               x8 : Bool;   // P2648.EPOS direct setpoint input/MDI positioning type
               x9 : Bool;   // P2651.EPOS direct setpoint input/MDI direction selection positive
               x10 : Bool;   // P2652.EPOS direct setpoint input/MDI direction selection negative
               x11 : Bool;   // Reserved
               x12 : Bool;   // P2649.EPOS direct setpoint input/MDI transfer type selection
               x13 : Bool;   // Reserved
               x14 : Bool;   // P2653.EPOS direct setpoint input/MDI setting-up selection
               x15 : Bool;   // P2647.EPOS direct setpoint input/MDI selection
               x0 : Bool;   // P2525.EPOS traversing block selection, bit 0
               x1 : Bool;   // P2526.EPOS traversing block selection, bit 1
               x2 : Bool;   // P2527.EPOS traversing block selection, bit 2
               x3 : Bool;   // P2528.EPOS traversing block selection, bit 3
               x4 : Bool;   // P2529.EPOS traversing block selection, bit 4
               x5 : Bool;   // P2530.EPOS traversing block selection, bit 5
               x6 : Bool;   // Reserved
               x7 : Bool;   // P2577.EPOS module correction activation
            END_STRUCT;
            tPOS_STW2 : Struct   // POSITIONER CONTROL WORD 3
               x8 : Bool;   // P2597.EPOS referencing type selection
               x9 : Bool;   // P2604.EPOS search for reference, start direction
               x10 : Bool;   // P2510.LR selecting measuring probe evaluation
               x11 : Bool;   // P2511.LR measuring probe evaluation edge
               x12 : Bool;   // Reserved
               x13 : Bool;   // Reserved
               x14 : Bool;   // P2582.EPOS software limit switch activation
               x15 : Bool;   // P2568.EPOS STOP cam activation
               x0 : Bool;   // P2655.EPOS select tracking mode
               x1 : Bool;   // P2596.EPOS set reference point
               x2 : Bool;   // P2612.EPOS search for reference cam
               x3 : Bool;   // Reserved
               x4 : Bool;   // Reserved
               x5 : Bool;   // P2591.EPOS jogging incremental
               x6 : Bool;   // Reserved
               x7 : Bool;   // Reserved
            END_STRUCT;
            iSTW2 : Int;   // P2045.CONTROL WORD 4
            iOVERRIDE : Int;   // P2646.Override % [0-16384]
            dMDI_TARPOS : DInt;   // P2642.Target position for MDI
            dMDI_VELOCITY : DInt;   // P2643.Speed reference for MDI
            iMDI_ACC : Int;   // P2644.Acceleration ramp % for MDI [0-16384]
            iMDI_DEC : Int;   // P2645.Deceleration ramp % for MDI [0-16384]
            iUser : Int;
         END_STRUCT;
      END_STRUCT;
   END_VAR
   VAR_TEMP
      TMP_dOldValue_AR1 : DInt;
      TMP_dOldValue_AR2 : DInt;
      TMP_x : Bool;
      TMP_i : Int;
      TMP_d : DInt;
      TMP_r : Real;
      TMP_a : ANY;
      TMP_dZero : DInt;
      TMP_xAlwaysON : Bool;
      TMP_rActualSpeed : Real;
      TMP_iAddressLength : Int;
      TMP_dActualPosMin_dmm : DInt;   // Actual position minimum tollerance [mm/10]
      TMP_dActualPosMax_dmm : DInt;   // Actual position maximum tollerance [mm/10]
      TMP_iRetVal : Int;
   END_VAR
   VAR_TEMP   // added for the SCL form of the ladder/FBD networks
      _w1 : Bool;
      _w2 : Bool;
      _w3 : Bool;
      _w4 : Bool;
      _w5 : Bool;
      _w6 : Bool;
      _w7 : Bool;
      _w8 : Bool;
      _w9 : Bool;
      _w10 : Bool;
      _w11 : Bool;
      _w12 : Bool;
   END_VAR
BEGIN

REGION Network 1 (STL): Save AR1 & AR2 value
   //    TAR1
   //    T     #TMP_dOldValue_AR1
   //    TAR2
   //    T     #TMP_dOldValue_AR2
END_REGION

REGION Network 2: #####_COSTANTS_#####
END_REGION

REGION Network 3 (STL): Initializing
         SET;
         S     #TMP_xAlwaysON;

         L     DINT#0;
         T     #TMP_dZero;

         CALL  FILL
         ( BVAL    := #TMP_dZero,
           RET_VAL := #TMP_iRetVal,
           BLK     := #STC_tPZD_Pos.tR
         );
END_REGION

REGION Network 4: #####_MOTOR_MODULE_#####
END_REGION

REGION Network 5 (STL): Check system data coerence
         L     #STC_tSYS_DATA.iIOAddress_MM;
         L     0;
         <I;
         L     10;
         JC    Err;

         L     #STC_tSYS_DATA.dMaxSpeed_rpm;
         L     DINT#0;
         <=D;
         L     11;
         JC    Err;

         L     #STC_tSYS_DATA.rK_rpm_mmMin;
         L     0.0;
         <=R;
         L     12;
         JC    Err;

         L     #STC_tSYS_DATA.rMaxAcc_m_s2;
         L     0.0;
         <=R;
         L     14;
         JC    Err;

         L     #STC_tSYS_DATA.rMaxDec_m_s2;
         L     0.0;
         <=R;
         L     15;
         JC    Err;

         L     12;
         T     #TMP_iAddressLength;

   //Compute destination position
         L;
         LAR1;
   //byte 1 = 10h (FIXED for S7)
         L     B#16#10;
         T     B[AR1, P#0.0];
   //byte 2 = data type
         L     B#16#4;  //4 = word
         T     B[AR1, P#1.0];
   //byte 3 & 4 = number of element
         L     #TMP_iAddressLength;  //Production data
         T     W[AR1, P#2.0];
   //byte 5 & 6 = number of DB
         L     0;  //DB production data
         T     W[AR1, P#4.0];
   //byte 7 = memory area
         L     B#16#81;  //81h = I (Input)
         T     B[AR1, P#6.0];
   //byte 8 & 9 = address. Bit 0,1,2 of tenth byte is bit offset
   //byte 7 = address (high). Valid value = 0-7. Bit 3,4,5,6,7 always 0

         L     #STC_tSYS_DATA.iIOAddress_MM;  //Item size
         SLW   3;
         T     W[AR1, P#8.0];
         SRD   16;
         AW    16#0007;
         T     B[AR1, P#7.0];

         CALL  BLKMOV
         ( SRCBLK  := #TMP_a,
           RET_VAL := #TMP_iRetVal,
           DSTBLK  := #STC_tPZD_Pos.tR
         );
END_REGION

REGION Network 6: #########################_POSITIONER_###########################
END_REGION

REGION Network 7: #####_MATCH_#####
END_REGION

REGION Network 8: Status signals
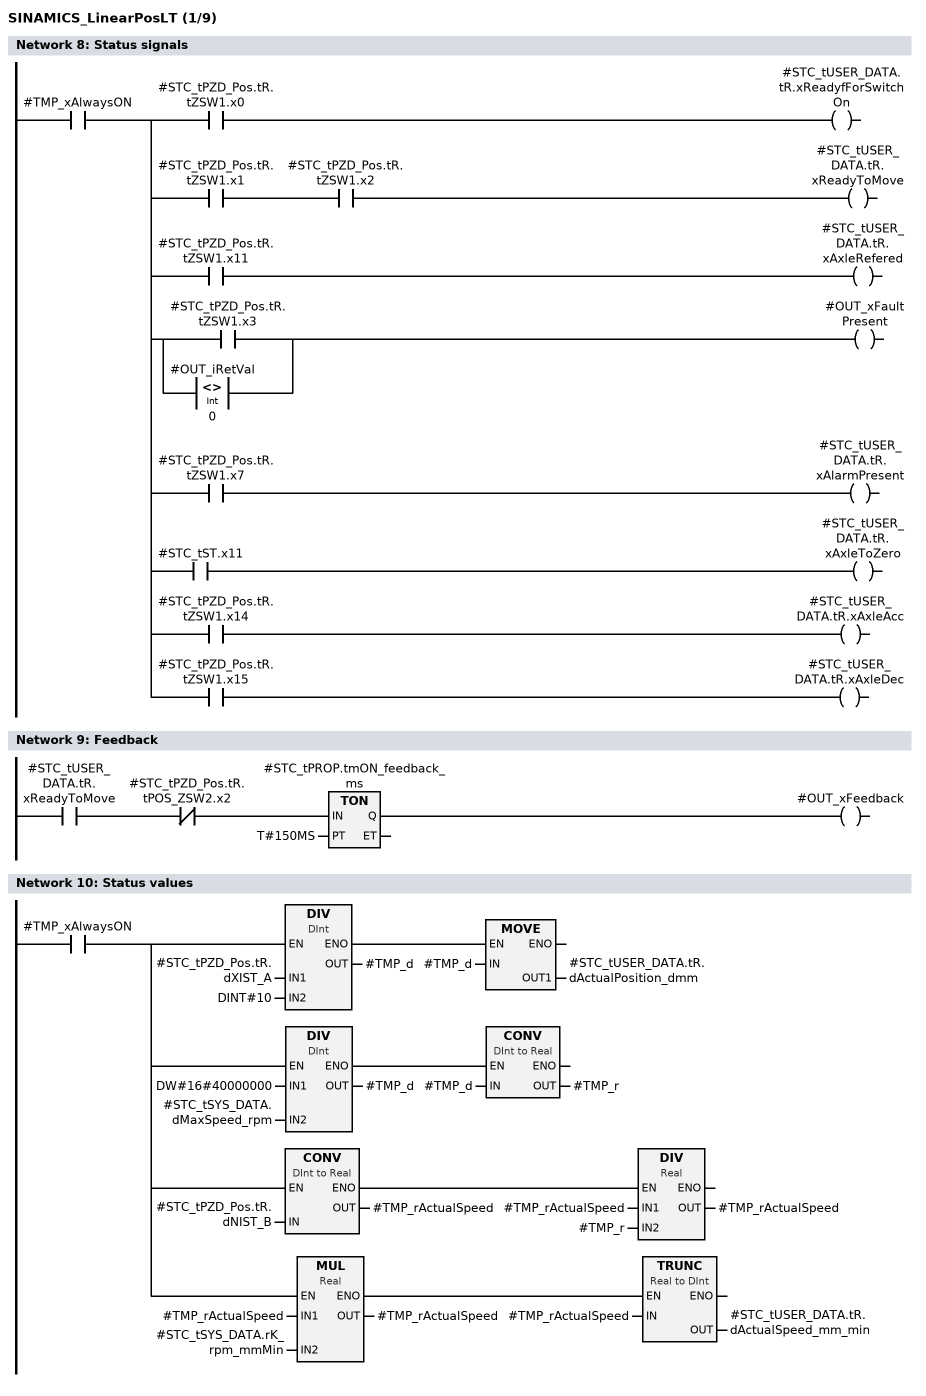
   RUNG wire#powerrail
      Contact( #TMP_xAlwaysON )
      wire#w1
      Contact( #STC_tPZD_Pos.tR.tZSW1.x0 )
      Coil( #STC_tUSER_DATA.tR.xReadyfForSwitchOn )
   END_RUNG
   RUNG wire#w1
      Contact( #STC_tPZD_Pos.tR.tZSW1.x1 )
      Contact( #STC_tPZD_Pos.tR.tZSW1.x2 )
      Coil( #STC_tUSER_DATA.tR.xReadyToMove )
   END_RUNG
   RUNG wire#w1
      Contact( #STC_tPZD_Pos.tR.tZSW1.x11 )
      Coil( #STC_tUSER_DATA.tR.xAxleRefered )
   END_RUNG
   RUNG wire#w1
      Contact( #STC_tPZD_Pos.tR.tZSW1.x3 )
      wire#w2
      Coil( #OUT_xFaultPresent )
   END_RUNG
   RUNG wire#w1
      { S7_Templates := "SrcType := Int" } NE_Contact(in1 := #OUT_iRetVal, in2 := 0)
   END_RUNG wire#w2
   RUNG wire#w1
      Contact( #STC_tPZD_Pos.tR.tZSW1.x7 )
      Coil( #STC_tUSER_DATA.tR.xAlarmPresent )
   END_RUNG
   RUNG wire#w1
      Contact( #STC_tST.x11 )
      Coil( #STC_tUSER_DATA.tR.xAxleToZero )
   END_RUNG
   RUNG wire#w1
      Contact( #STC_tPZD_Pos.tR.tZSW1.x14 )
      Coil( #STC_tUSER_DATA.tR.xAxleAcc )
   END_RUNG
   RUNG wire#w1
      Contact( #STC_tPZD_Pos.tR.tZSW1.x15 )
      Coil( #STC_tUSER_DATA.tR.xAxleDec )
   END_RUNG
   // the same network as SCL:
   #STC_tUSER_DATA.tR.xReadyfForSwitchOn := #TMP_xAlwaysON AND #STC_tPZD_Pos.tR.tZSW1.x0;
   #STC_tUSER_DATA.tR.xReadyToMove := #TMP_xAlwaysON AND #STC_tPZD_Pos.tR.tZSW1.x1 AND #STC_tPZD_Pos.tR.tZSW1.x2;
   #STC_tUSER_DATA.tR.xAxleRefered := #TMP_xAlwaysON AND #STC_tPZD_Pos.tR.tZSW1.x11;
   #OUT_xFaultPresent := #TMP_xAlwaysON AND (#STC_tPZD_Pos.tR.tZSW1.x3 OR (#OUT_iRetVal <> 0));
   #STC_tUSER_DATA.tR.xAlarmPresent := #TMP_xAlwaysON AND #STC_tPZD_Pos.tR.tZSW1.x7;
   #STC_tUSER_DATA.tR.xAxleToZero := #TMP_xAlwaysON AND #STC_tST.x11;
   #STC_tUSER_DATA.tR.xAxleAcc := #TMP_xAlwaysON AND #STC_tPZD_Pos.tR.tZSW1.x14;
   #STC_tUSER_DATA.tR.xAxleDec := #TMP_xAlwaysON AND #STC_tPZD_Pos.tR.tZSW1.x15;
END_REGION

REGION Network 9: Feedback
   #STC_tPROP.tmON_feedback_ms.TON(IN := #STC_tUSER_DATA.tR.xReadyToMove AND NOT #STC_tPZD_Pos.tR.tPOS_ZSW2.x2,
                           PT := T#150MS);
   #OUT_xFeedback := #STC_tPROP.tmON_feedback_ms.Q;
END_REGION

REGION Network 10: Status values
   RUNG wire#powerrail
      Contact( #TMP_xAlwaysON )
      wire#w1
      { S7_Templates := "SrcType := DInt"; S7_GenerateENO := "TRUE" } Div(in1 := #STC_tPZD_Pos.tR.dXIST_A, in2 := DINT#10, out => #TMP_d)
      { S7_GenerateENO := "TRUE" } Move(in := #TMP_d, out1 => #STC_tUSER_DATA.tR.dActualPosition_dmm)
   END_RUNG
   RUNG wire#w1
      { S7_Templates := "SrcType := DInt"; S7_GenerateENO := "TRUE" } Div(in1 := DW#16#40000000, in2 := #STC_tSYS_DATA.dMaxSpeed_rpm, out => #TMP_d)
      { S7_Templates := "[SrcType := DInt, DestType := Real]"; S7_GenerateENO := "TRUE" } Convert(in := #TMP_d, out => #TMP_r)
   END_RUNG
   RUNG wire#w1
      { S7_Templates := "[SrcType := DInt, DestType := Real]"; S7_GenerateENO := "TRUE" } Convert(in := #STC_tPZD_Pos.tR.dNIST_B, out => #TMP_rActualSpeed)
      { S7_Templates := "SrcType := Real"; S7_GenerateENO := "TRUE" } Div(in1 := #TMP_rActualSpeed, in2 := #TMP_r, out => #TMP_rActualSpeed)
   END_RUNG
   RUNG wire#w1
      { S7_Templates := "SrcType := Real"; S7_GenerateENO := "TRUE" } Mul(in1 := #TMP_rActualSpeed, in2 := #STC_tSYS_DATA.rK_rpm_mmMin, out => #TMP_rActualSpeed)
      { S7_Templates := "[SrcType := Real, DestType := DInt]"; S7_GenerateENO := "TRUE" } Trunc(in := #TMP_rActualSpeed, out => #STC_tUSER_DATA.tR.dActualSpeed_mm_min)
   END_RUNG
   // the same network as SCL:
   // ENO of a box is taken as its EN; it also drops when the box reports an error
   IF #TMP_xAlwaysON THEN
       #TMP_d := #STC_tPZD_Pos.tR.dXIST_A / DINT#10;
       #STC_tUSER_DATA.tR.dActualPosition_dmm := #TMP_d;
       #TMP_d := DW#16#40000000 / #STC_tSYS_DATA.dMaxSpeed_rpm;
       #TMP_r := DINT_TO_REAL(#TMP_d);
       #TMP_rActualSpeed := DINT_TO_REAL(#STC_tPZD_Pos.tR.dNIST_B);
       #TMP_rActualSpeed := #TMP_rActualSpeed / #TMP_r;
       #TMP_rActualSpeed := #TMP_rActualSpeed * #STC_tSYS_DATA.rK_rpm_mmMin;
       #STC_tUSER_DATA.tR.dActualSpeed_mm_min := TRUNC(#TMP_rActualSpeed);
   END_IF;
END_REGION

REGION Network 11: #####_STATUSES_#####
END_REGION

REGION Network 12: Type of positioning
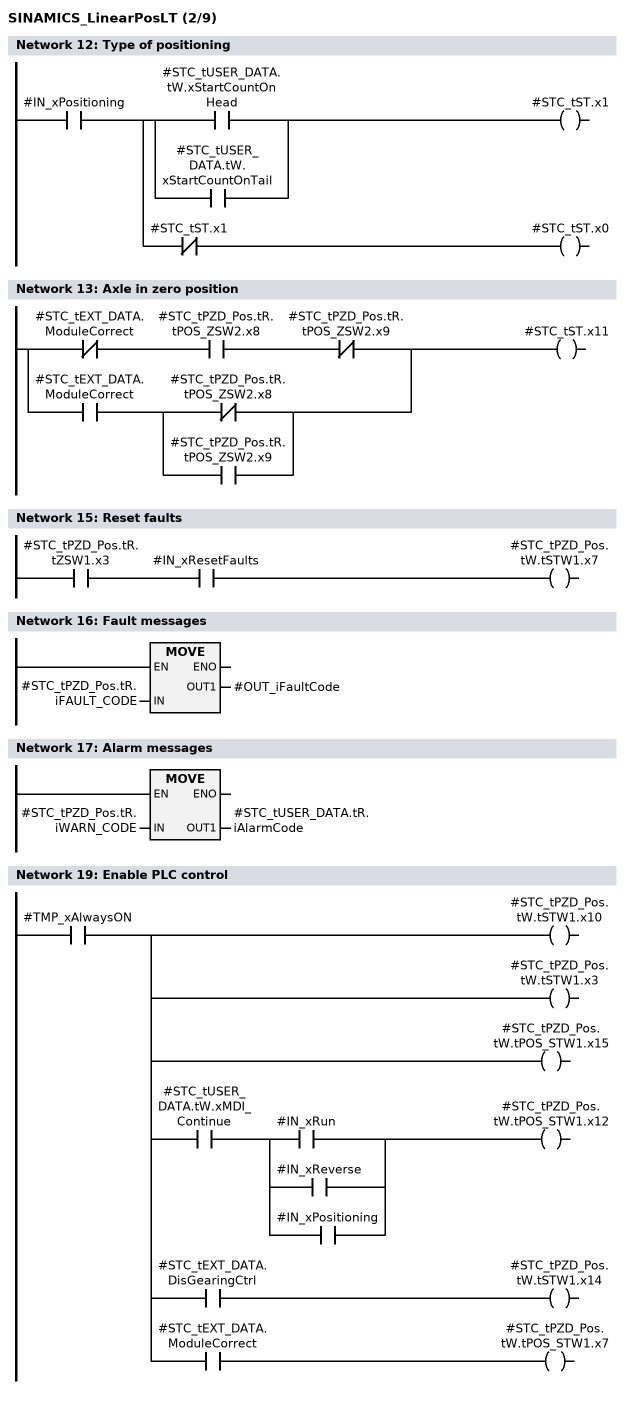
   RUNG wire#powerrail
      Contact( #IN_xPositioning )
      wire#w1
      Contact( #STC_tUSER_DATA.tW.xStartCountOnHead )
      wire#w2
      Coil( #STC_tST.x1 )
   END_RUNG
   RUNG wire#w1
      Contact( #STC_tUSER_DATA.tW.xStartCountOnTail )
   END_RUNG wire#w2
   RUNG wire#w1
      I_Contact( #STC_tST.x1 )
      Coil( #STC_tST.x0 )
   END_RUNG
   // the same network as SCL:
   #STC_tST.x1 := #IN_xPositioning AND (#STC_tUSER_DATA.tW.xStartCountOnHead OR #STC_tUSER_DATA.tW.xStartCountOnTail);
   #STC_tST.x0 := #IN_xPositioning AND NOT #STC_tST.x1;
END_REGION

REGION Network 13: Axle in zero position
   RUNG wire#powerrail
      I_Contact( #STC_tEXT_DATA.ModuleCorrect )
      Contact( #STC_tPZD_Pos.tR.tPOS_ZSW2.x8 )
      I_Contact( #STC_tPZD_Pos.tR.tPOS_ZSW2.x9 )
      wire#w1
      Coil( #STC_tST.x11 )
   END_RUNG
   RUNG wire#powerrail
      Contact( #STC_tEXT_DATA.ModuleCorrect )
      wire#w2
      I_Contact( #STC_tPZD_Pos.tR.tPOS_ZSW2.x8 )
   END_RUNG wire#w1
   RUNG wire#w2
      Contact( #STC_tPZD_Pos.tR.tPOS_ZSW2.x9 )
   END_RUNG wire#w1
   // the same network as SCL:
   #STC_tST.x11 := (NOT #STC_tEXT_DATA.ModuleCorrect AND #STC_tPZD_Pos.tR.tPOS_ZSW2.x8 AND NOT #STC_tPZD_Pos.tR.tPOS_ZSW2.x9) OR (#STC_tEXT_DATA.ModuleCorrect AND (NOT #STC_tPZD_Pos.tR.tPOS_ZSW2.x8 OR #STC_tPZD_Pos.tR.tPOS_ZSW2.x9));
END_REGION

REGION Network 14: #####_ALARMS_#####
END_REGION

REGION Network 15: Reset faults
   RUNG wire#powerrail
      Contact( #STC_tPZD_Pos.tR.tZSW1.x3 )
      Contact( #IN_xResetFaults )
      Coil( #STC_tPZD_Pos.tW.tSTW1.x7 )
   END_RUNG
   // the same network as SCL:
   #STC_tPZD_Pos.tW.tSTW1.x7 := #STC_tPZD_Pos.tR.tZSW1.x3 AND #IN_xResetFaults;
END_REGION

REGION Network 16: Fault messages
   RUNG wire#powerrail
      { S7_GenerateENO := "TRUE" } Move(in := #STC_tPZD_Pos.tR.iFAULT_CODE, out1 => #OUT_iFaultCode)
   END_RUNG
   // the same network as SCL:
   #OUT_iFaultCode := #STC_tPZD_Pos.tR.iFAULT_CODE;
END_REGION

REGION Network 17: Alarm messages
   RUNG wire#powerrail
      { S7_GenerateENO := "TRUE" } Move(in := #STC_tPZD_Pos.tR.iWARN_CODE, out1 => #STC_tUSER_DATA.tR.iAlarmCode)
   END_RUNG
   // the same network as SCL:
   #STC_tUSER_DATA.tR.iAlarmCode := #STC_tPZD_Pos.tR.iWARN_CODE;
END_REGION

REGION Network 18: #####_PHASES_&_LOGICS_#####
END_REGION

REGION Network 19: Enable PLC control
   RUNG wire#powerrail
      Contact( #TMP_xAlwaysON )
      wire#w1
      Coil( #STC_tPZD_Pos.tW.tSTW1.x10 )
   END_RUNG
   RUNG wire#w1
      Coil( #STC_tPZD_Pos.tW.tSTW1.x3 )
   END_RUNG
   RUNG wire#w1
      Coil( #STC_tPZD_Pos.tW.tPOS_STW1.x15 )
   END_RUNG
   RUNG wire#w1
      Contact( #STC_tUSER_DATA.tW.xMDI_Continue )
      wire#w2
      Contact( #IN_xRun )
      wire#w3
      Coil( #STC_tPZD_Pos.tW.tPOS_STW1.x12 )
   END_RUNG
   RUNG wire#w2
      Contact( #IN_xReverse )
   END_RUNG wire#w3
   RUNG wire#w2
      Contact( #IN_xPositioning )
   END_RUNG wire#w3
   RUNG wire#w1
      Contact( #STC_tEXT_DATA.DisGearingCtrl )
      Coil( #STC_tPZD_Pos.tW.tSTW1.x14 )
   END_RUNG
   RUNG wire#w1
      Contact( #STC_tEXT_DATA.ModuleCorrect )
      Coil( #STC_tPZD_Pos.tW.tPOS_STW1.x7 )
   END_RUNG
   // the same network as SCL:
   #STC_tPZD_Pos.tW.tSTW1.x10 := #TMP_xAlwaysON;
   #STC_tPZD_Pos.tW.tSTW1.x3 := #TMP_xAlwaysON;
   #STC_tPZD_Pos.tW.tPOS_STW1.x15 := #TMP_xAlwaysON;
   #STC_tPZD_Pos.tW.tPOS_STW1.x12 := #TMP_xAlwaysON AND #STC_tUSER_DATA.tW.xMDI_Continue AND (#IN_xRun OR #IN_xReverse OR #IN_xPositioning);
   #STC_tPZD_Pos.tW.tSTW1.x14 := #TMP_xAlwaysON AND #STC_tEXT_DATA.DisGearingCtrl;
   #STC_tPZD_Pos.tW.tPOS_STW1.x7 := #TMP_xAlwaysON AND #STC_tEXT_DATA.ModuleCorrect;
END_REGION

REGION Network 20: Drive Enable
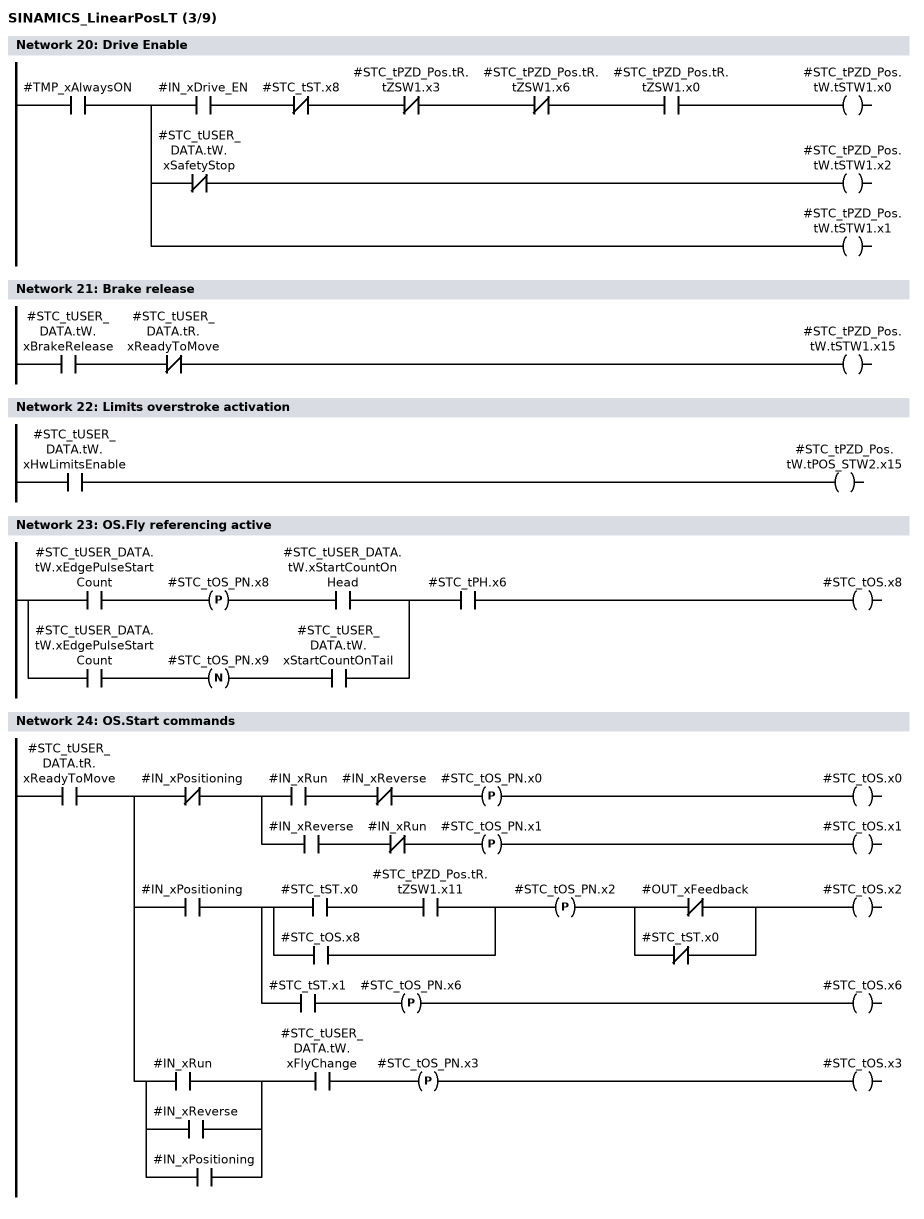
   RUNG wire#powerrail
      Contact( #TMP_xAlwaysON )
      wire#w1
      Contact( #IN_xDrive_EN )
      I_Contact( #STC_tST.x8 )
      I_Contact( #STC_tPZD_Pos.tR.tZSW1.x3 )
      I_Contact( #STC_tPZD_Pos.tR.tZSW1.x6 )
      Contact( #STC_tPZD_Pos.tR.tZSW1.x0 )
      Coil( #STC_tPZD_Pos.tW.tSTW1.x0 )
   END_RUNG
   RUNG wire#w1
      I_Contact( #STC_tUSER_DATA.tW.xSafetyStop )
      Coil( #STC_tPZD_Pos.tW.tSTW1.x2 )
   END_RUNG
   RUNG wire#w1
      Coil( #STC_tPZD_Pos.tW.tSTW1.x1 )
   END_RUNG
   // the same network as SCL:
   #STC_tPZD_Pos.tW.tSTW1.x0 := #TMP_xAlwaysON AND #IN_xDrive_EN AND NOT #STC_tST.x8 AND NOT #STC_tPZD_Pos.tR.tZSW1.x3 AND NOT #STC_tPZD_Pos.tR.tZSW1.x6 AND #STC_tPZD_Pos.tR.tZSW1.x0;
   #STC_tPZD_Pos.tW.tSTW1.x2 := #TMP_xAlwaysON AND NOT #STC_tUSER_DATA.tW.xSafetyStop;
   #STC_tPZD_Pos.tW.tSTW1.x1 := #TMP_xAlwaysON;
END_REGION

REGION Network 21: Brake release
   RUNG wire#powerrail
      Contact( #STC_tUSER_DATA.tW.xBrakeRelease )
      I_Contact( #STC_tUSER_DATA.tR.xReadyToMove )
      Coil( #STC_tPZD_Pos.tW.tSTW1.x15 )
   END_RUNG
   // the same network as SCL:
   #STC_tPZD_Pos.tW.tSTW1.x15 := #STC_tUSER_DATA.tW.xBrakeRelease AND NOT #STC_tUSER_DATA.tR.xReadyToMove;
END_REGION

REGION Network 22: Limits overstroke activation
   RUNG wire#powerrail
      Contact( #STC_tUSER_DATA.tW.xHwLimitsEnable )
      Coil( #STC_tPZD_Pos.tW.tPOS_STW2.x15 )
   END_RUNG
   // the same network as SCL:
   #STC_tPZD_Pos.tW.tPOS_STW2.x15 := #STC_tUSER_DATA.tW.xHwLimitsEnable;
END_REGION

REGION Network 23: OS.Fly referencing active
   RUNG wire#powerrail
      Contact( #STC_tUSER_DATA.tW.xEdgePulseStartCount )
      P_Trig( #STC_tOS_PN.x8 )
      Contact( #STC_tUSER_DATA.tW.xStartCountOnHead )
      wire#w1
      Contact( #STC_tPH.x6 )
      Coil( #STC_tOS.x8 )
   END_RUNG
   RUNG wire#powerrail
      Contact( #STC_tUSER_DATA.tW.xEdgePulseStartCount )
      N_Trig( #STC_tOS_PN.x9 )
      Contact( #STC_tUSER_DATA.tW.xStartCountOnTail )
   END_RUNG wire#w1
   // the same network as SCL:
   #_w1 := #STC_tUSER_DATA.tW.xEdgePulseStartCount AND NOT #STC_tOS_PN.x8;   // rising edge
   #STC_tOS_PN.x8 := #STC_tUSER_DATA.tW.xEdgePulseStartCount;
   #_w2 := NOT #STC_tUSER_DATA.tW.xEdgePulseStartCount AND #STC_tOS_PN.x9;   // falling edge
   #STC_tOS_PN.x9 := #STC_tUSER_DATA.tW.xEdgePulseStartCount;
   #STC_tOS.x8 := ((#_w1 AND #STC_tUSER_DATA.tW.xStartCountOnHead) OR (#_w2 AND #STC_tUSER_DATA.tW.xStartCountOnTail)) AND #STC_tPH.x6;
END_REGION

REGION Network 24: OS.Start commands
   RUNG wire#powerrail
      Contact( #STC_tUSER_DATA.tR.xReadyToMove )
      wire#w1
      I_Contact( #IN_xPositioning )
      wire#w2
      Contact( #IN_xRun )
      I_Contact( #IN_xReverse )
      P_Trig( #STC_tOS_PN.x0 )
      Coil( #STC_tOS.x0 )
   END_RUNG
   RUNG wire#w2
      Contact( #IN_xReverse )
      I_Contact( #IN_xRun )
      P_Trig( #STC_tOS_PN.x1 )
      Coil( #STC_tOS.x1 )
   END_RUNG
   RUNG wire#w1
      Contact( #IN_xPositioning )
      wire#w3
      Contact( #STC_tST.x0 )
      Contact( #STC_tPZD_Pos.tR.tZSW1.x11 )
      wire#w4
      P_Trig( #STC_tOS_PN.x2 )
      wire#w5
      I_Contact( #OUT_xFeedback )
      wire#w6
      Coil( #STC_tOS.x2 )
   END_RUNG
   RUNG wire#w3
      Contact( #STC_tOS.x8 )
   END_RUNG wire#w4
   RUNG wire#w5
      I_Contact( #STC_tST.x0 )
   END_RUNG wire#w6
   RUNG wire#w3
      Contact( #STC_tST.x1 )
      P_Trig( #STC_tOS_PN.x6 )
      Coil( #STC_tOS.x6 )
   END_RUNG
   RUNG wire#w1
      Contact( #IN_xRun )
      wire#w7
      Contact( #STC_tUSER_DATA.tW.xFlyChange )
      P_Trig( #STC_tOS_PN.x3 )
      Coil( #STC_tOS.x3 )
   END_RUNG
   RUNG wire#w1
      Contact( #IN_xReverse )
   END_RUNG wire#w7
   RUNG wire#w1
      Contact( #IN_xPositioning )
   END_RUNG wire#w7
   // the same network as SCL:
   #_w1 := #STC_tUSER_DATA.tR.xReadyToMove AND NOT #IN_xPositioning;
   #_w2 := #_w1 AND #IN_xRun AND NOT #IN_xReverse;
   #_w3 := #_w2 AND NOT #STC_tOS_PN.x0;   // rising edge
   #STC_tOS_PN.x0 := #_w2;
   #STC_tOS.x0 := #_w3;
   #_w4 := #_w1 AND #IN_xReverse AND NOT #IN_xRun;
   #_w5 := #_w4 AND NOT #STC_tOS_PN.x1;   // rising edge
   #STC_tOS_PN.x1 := #_w4;
   #STC_tOS.x1 := #_w5;
   #_w6 := #STC_tUSER_DATA.tR.xReadyToMove AND #IN_xPositioning;
   #_w7 := #_w6 AND ((#STC_tST.x0 AND #STC_tPZD_Pos.tR.tZSW1.x11) OR #STC_tOS.x8);
   #_w8 := #_w7 AND NOT #STC_tOS_PN.x2;   // rising edge
   #STC_tOS_PN.x2 := #_w7;
   #STC_tOS.x2 := #_w8 AND (NOT #OUT_xFeedback OR NOT #STC_tST.x0);
   #_w9 := #_w6 AND #STC_tST.x1;
   #_w10 := #_w9 AND NOT #STC_tOS_PN.x6;   // rising edge
   #STC_tOS_PN.x6 := #_w9;
   #STC_tOS.x6 := #_w10;
   #_w11 := #STC_tUSER_DATA.tR.xReadyToMove AND (#IN_xRun OR #IN_xReverse OR #IN_xPositioning) AND #STC_tUSER_DATA.tW.xFlyChange;
   #_w12 := #_w11 AND NOT #STC_tOS_PN.x3;   // rising edge
   #STC_tOS_PN.x3 := #_w11;
   #STC_tOS.x3 := #_w12;
END_REGION

REGION Network 25: Sending data copy
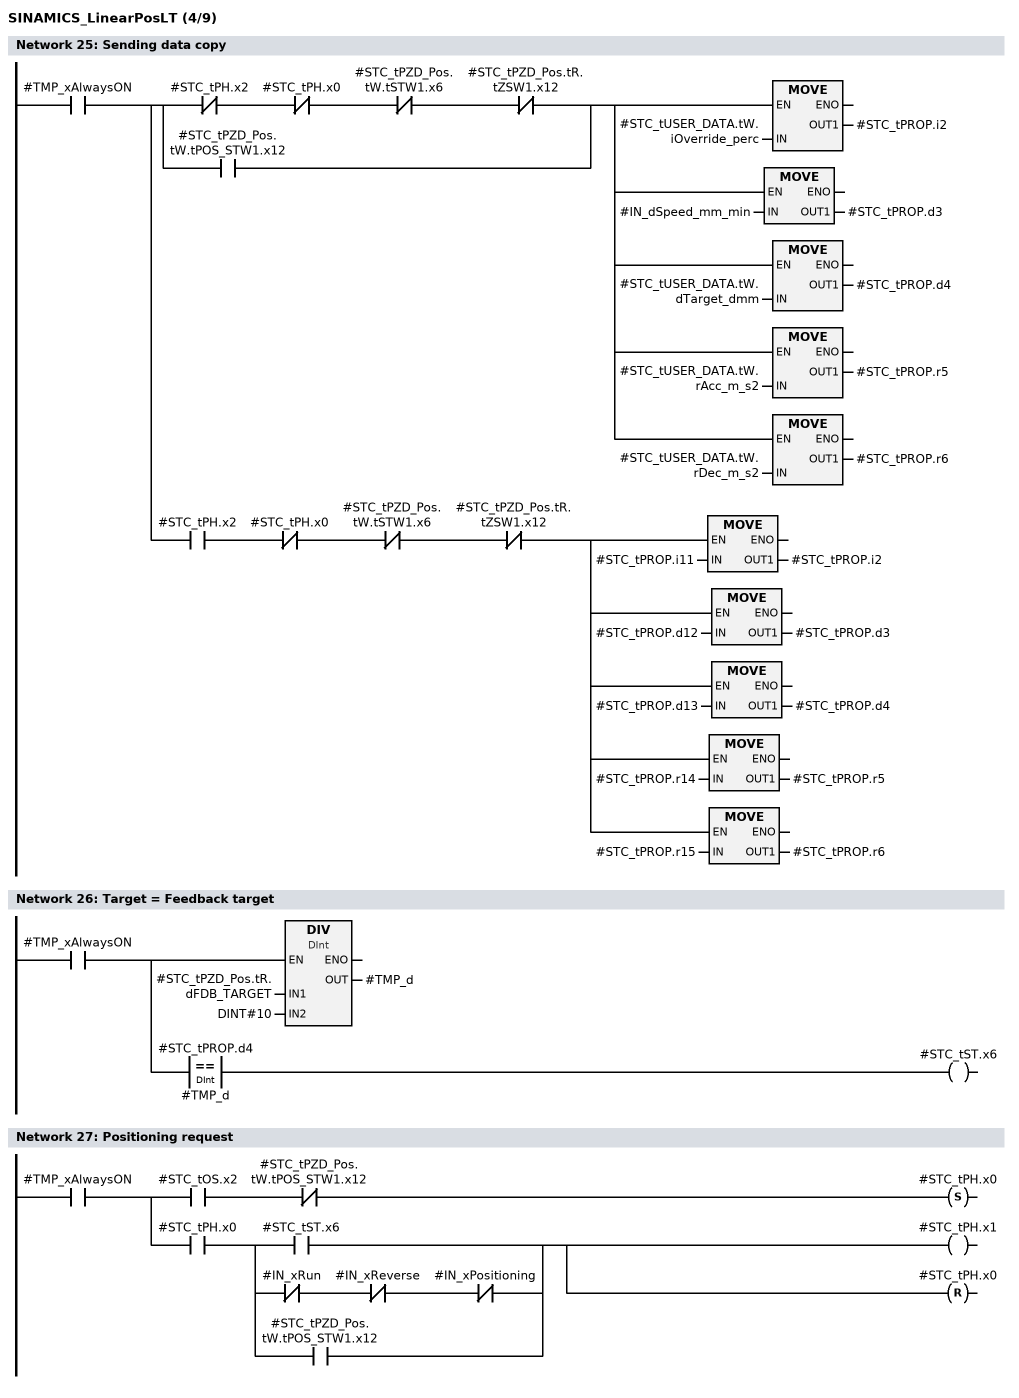
   RUNG wire#powerrail
      Contact( #TMP_xAlwaysON )
      wire#w1
      I_Contact( #STC_tPH.x2 )
      I_Contact( #STC_tPH.x0 )
      I_Contact( #STC_tPZD_Pos.tW.tSTW1.x6 )
      I_Contact( #STC_tPZD_Pos.tR.tZSW1.x12 )
      wire#w2
      { S7_GenerateENO := "TRUE" } Move(in := #STC_tUSER_DATA.tW.iOverride_perc, out1 => #STC_tPROP.i2)
   END_RUNG
   RUNG wire#w1
      Contact( #STC_tPZD_Pos.tW.tPOS_STW1.x12 )
   END_RUNG wire#w2
   RUNG wire#w2
      { S7_GenerateENO := "TRUE" } Move(in := #IN_dSpeed_mm_min, out1 => #STC_tPROP.d3)
   END_RUNG
   RUNG wire#w2
      { S7_GenerateENO := "TRUE" } Move(in := #STC_tUSER_DATA.tW.dTarget_dmm, out1 => #STC_tPROP.d4)
   END_RUNG
   RUNG wire#w2
      { S7_GenerateENO := "TRUE" } Move(in := #STC_tUSER_DATA.tW.rAcc_m_s2, out1 => #STC_tPROP.r5)
   END_RUNG
   RUNG wire#w2
      { S7_GenerateENO := "TRUE" } Move(in := #STC_tUSER_DATA.tW.rDec_m_s2, out1 => #STC_tPROP.r6)
   END_RUNG
   RUNG wire#w1
      Contact( #STC_tPH.x2 )
      I_Contact( #STC_tPH.x0 )
      I_Contact( #STC_tPZD_Pos.tW.tSTW1.x6 )
      I_Contact( #STC_tPZD_Pos.tR.tZSW1.x12 )
      wire#w3
      { S7_GenerateENO := "TRUE" } Move(in := #STC_tPROP.i11, out1 => #STC_tPROP.i2)
   END_RUNG
   RUNG wire#w3
      { S7_GenerateENO := "TRUE" } Move(in := #STC_tPROP.d12, out1 => #STC_tPROP.d3)
   END_RUNG
   RUNG wire#w3
      { S7_GenerateENO := "TRUE" } Move(in := #STC_tPROP.d13, out1 => #STC_tPROP.d4)
   END_RUNG
   RUNG wire#w3
      { S7_GenerateENO := "TRUE" } Move(in := #STC_tPROP.r14, out1 => #STC_tPROP.r5)
   END_RUNG
   RUNG wire#w3
      { S7_GenerateENO := "TRUE" } Move(in := #STC_tPROP.r15, out1 => #STC_tPROP.r6)
   END_RUNG
   // the same network as SCL:
   IF #TMP_xAlwaysON AND ((NOT #STC_tPH.x2 AND NOT #STC_tPH.x0 AND NOT #STC_tPZD_Pos.tW.tSTW1.x6 AND NOT #STC_tPZD_Pos.tR.tZSW1.x12) OR #STC_tPZD_Pos.tW.tPOS_STW1.x12) THEN
       #STC_tPROP.i2 := #STC_tUSER_DATA.tW.iOverride_perc;
       #STC_tPROP.d3 := #IN_dSpeed_mm_min;
       #STC_tPROP.d4 := #STC_tUSER_DATA.tW.dTarget_dmm;
       #STC_tPROP.r5 := #STC_tUSER_DATA.tW.rAcc_m_s2;
       #STC_tPROP.r6 := #STC_tUSER_DATA.tW.rDec_m_s2;
   END_IF;
   IF #TMP_xAlwaysON AND #STC_tPH.x2 AND NOT #STC_tPH.x0 AND NOT #STC_tPZD_Pos.tW.tSTW1.x6 AND NOT #STC_tPZD_Pos.tR.tZSW1.x12 THEN
       #STC_tPROP.i2 := #STC_tPROP.i11;
       #STC_tPROP.d3 := #STC_tPROP.d12;
       #STC_tPROP.d4 := #STC_tPROP.d13;
       #STC_tPROP.r5 := #STC_tPROP.r14;
       #STC_tPROP.r6 := #STC_tPROP.r15;
   END_IF;
END_REGION

REGION Network 26: Target = Feedback target
   RUNG wire#powerrail
      Contact( #TMP_xAlwaysON )
      wire#w1
      { S7_Templates := "SrcType := DInt"; S7_GenerateENO := "TRUE" } Div(in1 := #STC_tPZD_Pos.tR.dFDB_TARGET, in2 := DINT#10, out => #TMP_d)
   END_RUNG
   RUNG wire#w1
      { S7_Templates := "SrcType := DInt" } EQ_Contact(in1 := #STC_tPROP.d4, in2 := #TMP_d)
      Coil( #STC_tST.x6 )
   END_RUNG
   // the same network as SCL:
   IF #TMP_xAlwaysON THEN #TMP_d := #STC_tPZD_Pos.tR.dFDB_TARGET / DINT#10; END_IF;
   #STC_tST.x6 := #TMP_xAlwaysON AND (#STC_tPROP.d4 = #TMP_d);
END_REGION

REGION Network 27: Positioning request
   RUNG wire#powerrail
      Contact( #TMP_xAlwaysON )
      wire#w1
      Contact( #STC_tOS.x2 )
      I_Contact( #STC_tPZD_Pos.tW.tPOS_STW1.x12 )
      S_Coil( #STC_tPH.x0 )
   END_RUNG
   RUNG wire#w1
      Contact( #STC_tPH.x0 )
      wire#w2
      Contact( #STC_tST.x6 )
      wire#w3
      Coil( #STC_tPH.x1 )
   END_RUNG
   RUNG wire#w2
      I_Contact( #IN_xRun )
      I_Contact( #IN_xReverse )
      I_Contact( #IN_xPositioning )
   END_RUNG wire#w3
   RUNG wire#w2
      Contact( #STC_tPZD_Pos.tW.tPOS_STW1.x12 )
   END_RUNG wire#w3
   RUNG wire#w3
      R_Coil( #STC_tPH.x0 )
   END_RUNG
   // the same network as SCL:
   IF #TMP_xAlwaysON AND #STC_tOS.x2 AND NOT #STC_tPZD_Pos.tW.tPOS_STW1.x12 THEN #STC_tPH.x0 := TRUE; END_IF;
   #STC_tPH.x1 := #TMP_xAlwaysON AND #STC_tPH.x0 AND (#STC_tST.x6 OR (NOT #IN_xRun AND NOT #IN_xReverse AND NOT #IN_xPositioning) OR #STC_tPZD_Pos.tW.tPOS_STW1.x12);
   IF #STC_tPH.x1 THEN #STC_tPH.x0 := FALSE; END_IF;
END_REGION

REGION Network 28: Fly change request
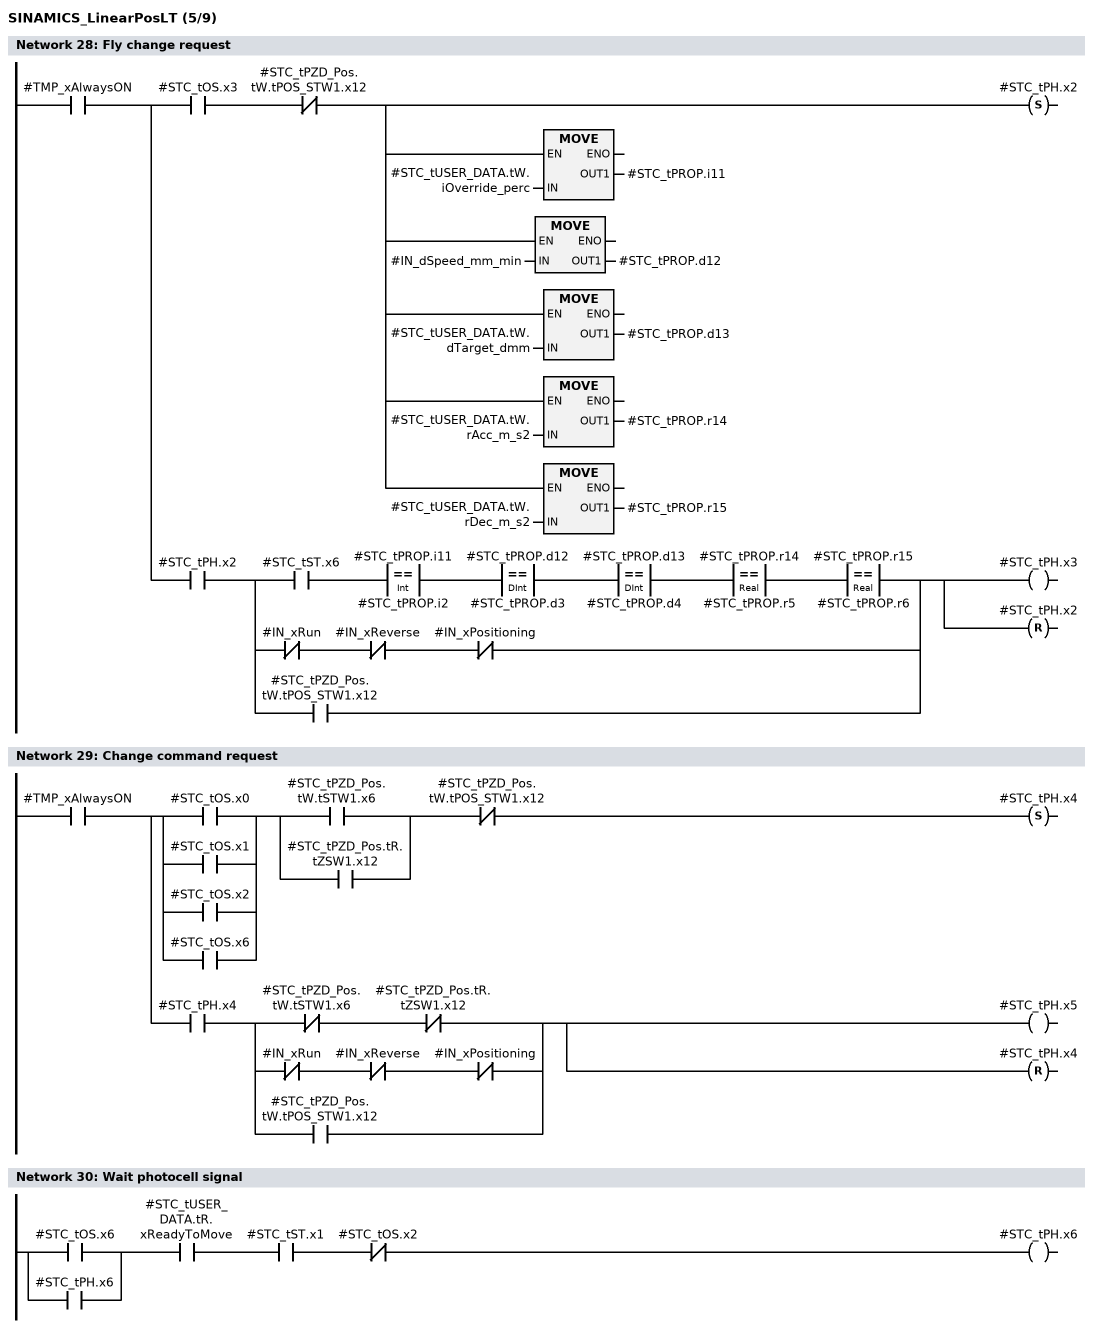
   RUNG wire#powerrail
      Contact( #TMP_xAlwaysON )
      wire#w1
      Contact( #STC_tOS.x3 )
      I_Contact( #STC_tPZD_Pos.tW.tPOS_STW1.x12 )
      wire#w2
      S_Coil( #STC_tPH.x2 )
   END_RUNG
   RUNG wire#w2
      Move(in := #STC_tUSER_DATA.tW.iOverride_perc, out1 => #STC_tPROP.i11)
   END_RUNG
   RUNG wire#w2
      Move(in := #IN_dSpeed_mm_min, out1 => #STC_tPROP.d12)
   END_RUNG
   RUNG wire#w2
      Move(in := #STC_tUSER_DATA.tW.dTarget_dmm, out1 => #STC_tPROP.d13)
   END_RUNG
   RUNG wire#w2
      Move(in := #STC_tUSER_DATA.tW.rAcc_m_s2, out1 => #STC_tPROP.r14)
   END_RUNG
   RUNG wire#w2
      Move(in := #STC_tUSER_DATA.tW.rDec_m_s2, out1 => #STC_tPROP.r15)
   END_RUNG
   RUNG wire#w1
      Contact( #STC_tPH.x2 )
      wire#w3
      Contact( #STC_tST.x6 )
      { S7_Templates := "SrcType := Int" } EQ_Contact(in1 := #STC_tPROP.i11, in2 := #STC_tPROP.i2)
      { S7_Templates := "SrcType := DInt" } EQ_Contact(in1 := #STC_tPROP.d12, in2 := #STC_tPROP.d3)
      { S7_Templates := "SrcType := DInt" } EQ_Contact(in1 := #STC_tPROP.d13, in2 := #STC_tPROP.d4)
      { S7_Templates := "SrcType := Real" } EQ_Contact(in1 := #STC_tPROP.r14, in2 := #STC_tPROP.r5)
      { S7_Templates := "SrcType := Real" } EQ_Contact(in1 := #STC_tPROP.r15, in2 := #STC_tPROP.r6)
      wire#w4
      Coil( #STC_tPH.x3 )
   END_RUNG
   RUNG wire#w3
      I_Contact( #IN_xRun )
      I_Contact( #IN_xReverse )
      I_Contact( #IN_xPositioning )
   END_RUNG wire#w4
   RUNG wire#w3
      Contact( #STC_tPZD_Pos.tW.tPOS_STW1.x12 )
   END_RUNG wire#w4
   RUNG wire#w4
      R_Coil( #STC_tPH.x2 )
   END_RUNG
   // the same network as SCL:
   IF #TMP_xAlwaysON AND #STC_tOS.x3 AND NOT #STC_tPZD_Pos.tW.tPOS_STW1.x12 THEN
       #STC_tPH.x2 := TRUE;
       #STC_tPROP.i11 := #STC_tUSER_DATA.tW.iOverride_perc;
       #STC_tPROP.d12 := #IN_dSpeed_mm_min;
       #STC_tPROP.d13 := #STC_tUSER_DATA.tW.dTarget_dmm;
       #STC_tPROP.r14 := #STC_tUSER_DATA.tW.rAcc_m_s2;
       #STC_tPROP.r15 := #STC_tUSER_DATA.tW.rDec_m_s2;
   END_IF;
   #STC_tPH.x3 := #TMP_xAlwaysON AND #STC_tPH.x2 AND ((#STC_tST.x6 AND (#STC_tPROP.i11 = #STC_tPROP.i2) AND (#STC_tPROP.d12 = #STC_tPROP.d3) AND (#STC_tPROP.d13 = #STC_tPROP.d4) AND (#STC_tPROP.r14 = #STC_tPROP.r5) AND (#STC_tPROP.r15 = #STC_tPROP.r6)) OR (NOT #IN_xRun AND NOT #IN_xReverse AND NOT #IN_xPositioning) OR #STC_tPZD_Pos.tW.tPOS_STW1.x12);
   IF #STC_tPH.x3 THEN #STC_tPH.x2 := FALSE; END_IF;
END_REGION

REGION Network 29: Change command request
   RUNG wire#powerrail
      Contact( #TMP_xAlwaysON )
      wire#w1
      Contact( #STC_tOS.x0 )
      wire#w2
      Contact( #STC_tPZD_Pos.tW.tSTW1.x6 )
      wire#w3
      I_Contact( #STC_tPZD_Pos.tW.tPOS_STW1.x12 )
      S_Coil( #STC_tPH.x4 )
   END_RUNG
   RUNG wire#w1
      Contact( #STC_tOS.x1 )
   END_RUNG wire#w2
   RUNG wire#w1
      Contact( #STC_tOS.x2 )
   END_RUNG wire#w2
   RUNG wire#w1
      Contact( #STC_tOS.x6 )
   END_RUNG wire#w2
   RUNG wire#w2
      Contact( #STC_tPZD_Pos.tR.tZSW1.x12 )
   END_RUNG wire#w3
   RUNG wire#w1
      Contact( #STC_tPH.x4 )
      wire#w4
      I_Contact( #STC_tPZD_Pos.tW.tSTW1.x6 )
      I_Contact( #STC_tPZD_Pos.tR.tZSW1.x12 )
      wire#w5
      Coil( #STC_tPH.x5 )
   END_RUNG
   RUNG wire#w4
      I_Contact( #IN_xRun )
      I_Contact( #IN_xReverse )
      I_Contact( #IN_xPositioning )
   END_RUNG wire#w5
   RUNG wire#w4
      Contact( #STC_tPZD_Pos.tW.tPOS_STW1.x12 )
   END_RUNG wire#w5
   RUNG wire#w5
      R_Coil( #STC_tPH.x4 )
   END_RUNG
   // the same network as SCL:
   IF #TMP_xAlwaysON AND (#STC_tOS.x0 OR #STC_tOS.x1 OR #STC_tOS.x2 OR #STC_tOS.x6) AND (#STC_tPZD_Pos.tW.tSTW1.x6 OR #STC_tPZD_Pos.tR.tZSW1.x12) AND NOT #STC_tPZD_Pos.tW.tPOS_STW1.x12 THEN
       #STC_tPH.x4 := TRUE;
   END_IF;
   #STC_tPH.x5 := #TMP_xAlwaysON AND #STC_tPH.x4 AND ((NOT #STC_tPZD_Pos.tW.tSTW1.x6 AND NOT #STC_tPZD_Pos.tR.tZSW1.x12) OR (NOT #IN_xRun AND NOT #IN_xReverse AND NOT #IN_xPositioning) OR #STC_tPZD_Pos.tW.tPOS_STW1.x12);
   IF #STC_tPH.x5 THEN #STC_tPH.x4 := FALSE; END_IF;
END_REGION

REGION Network 30: Wait photocell signal
   RUNG wire#powerrail
      Contact( #STC_tOS.x6 )
      wire#w1
      Contact( #STC_tUSER_DATA.tR.xReadyToMove )
      Contact( #STC_tST.x1 )
      I_Contact( #STC_tOS.x2 )
      Coil( #STC_tPH.x6 )
   END_RUNG
   RUNG wire#powerrail
      Contact( #STC_tPH.x6 )
   END_RUNG wire#w1
   // the same network as SCL:
   #STC_tPH.x6 := (#STC_tOS.x6 OR #STC_tPH.x6) AND #STC_tUSER_DATA.tR.xReadyToMove AND #STC_tST.x1 AND NOT #STC_tOS.x2;
END_REGION

REGION Network 31: Run/Reverse Commands
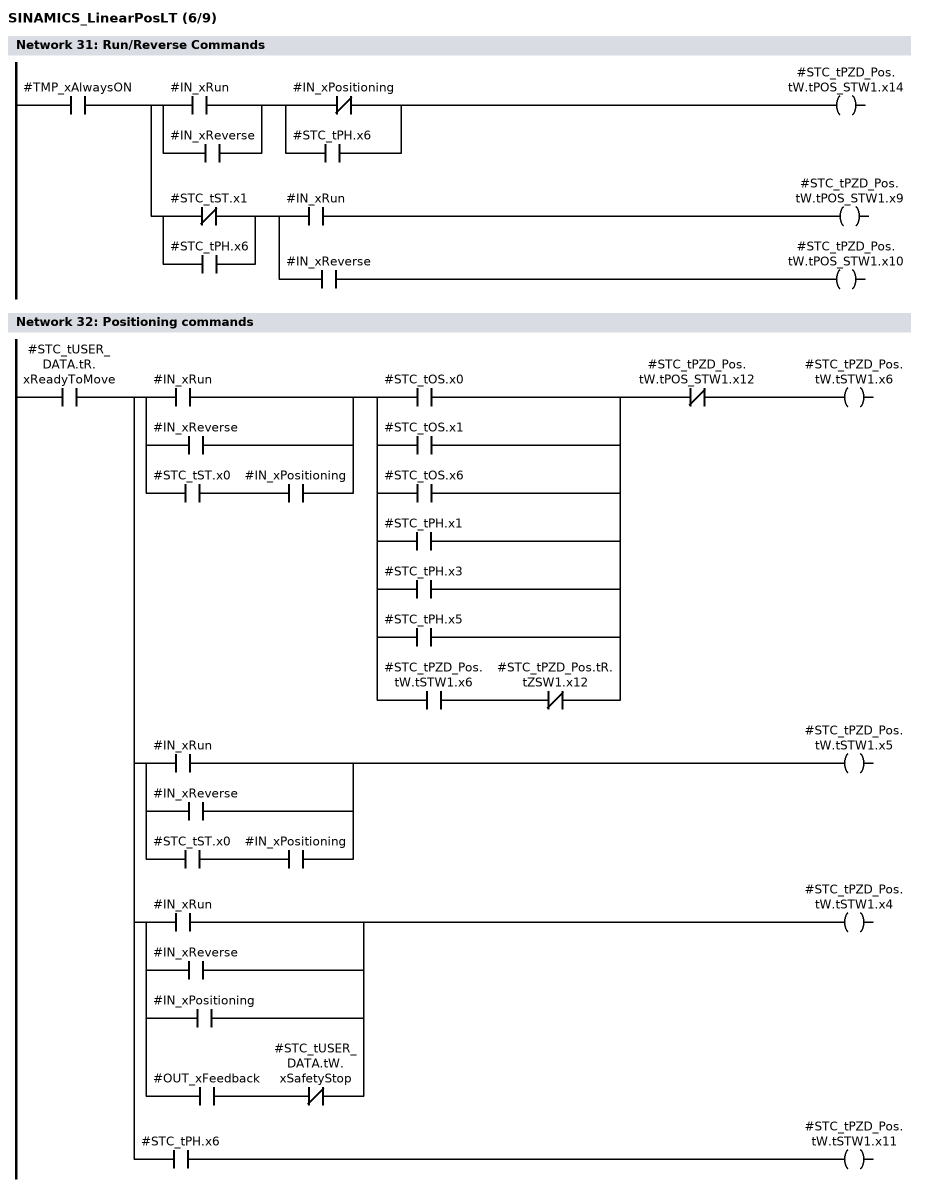
   RUNG wire#powerrail
      Contact( #TMP_xAlwaysON )
      wire#w1
      Contact( #IN_xRun )
      wire#w2
      I_Contact( #IN_xPositioning )
      wire#w3
      Coil( #STC_tPZD_Pos.tW.tPOS_STW1.x14 )
   END_RUNG
   RUNG wire#w1
      Contact( #IN_xReverse )
   END_RUNG wire#w2
   RUNG wire#w2
      Contact( #STC_tPH.x6 )
   END_RUNG wire#w3
   RUNG wire#w1
      I_Contact( #STC_tST.x1 )
      wire#w4
      Contact( #IN_xRun )
      Coil( #STC_tPZD_Pos.tW.tPOS_STW1.x9 )
   END_RUNG
   RUNG wire#w1
      Contact( #STC_tPH.x6 )
   END_RUNG wire#w4
   RUNG wire#w4
      Contact( #IN_xReverse )
      Coil( #STC_tPZD_Pos.tW.tPOS_STW1.x10 )
   END_RUNG
   // the same network as SCL:
   #STC_tPZD_Pos.tW.tPOS_STW1.x14 := #TMP_xAlwaysON AND (#IN_xRun OR #IN_xReverse) AND (NOT #IN_xPositioning OR #STC_tPH.x6);
   #_w1 := #TMP_xAlwaysON AND (NOT #STC_tST.x1 OR #STC_tPH.x6);
   #STC_tPZD_Pos.tW.tPOS_STW1.x9 := #_w1 AND #IN_xRun;
   #STC_tPZD_Pos.tW.tPOS_STW1.x10 := #_w1 AND #IN_xReverse;
END_REGION

